// TIA Portal project "XSFW_TIA31001_B0_V15.1" (V15.1)

(* hardware
DEVICE "S7-1200 station_1"  S7-1200 Station
   slot 0: "Rack_0"  S7-1200 Rack  Rack  V1.0
   slot 1: "PLC_Divider"  CPU 1214C DC/DC/DC  6ES7 214-1AG40-0XB0  V4.2
   slot 2: "DI 16/DQ 16x24VDC_1"  6ES7 223-1BL32-0XB0  V2.0
   slot 3: "AI 4x13BIT/AQ 2x14BIT_1"  6ES7 234-4HE32-0XB0  V2.0
   slot 101: "CM 1242-5"  CM 1242-5  6GK7 242-5DX30-0XE0  V1.0
DEVICE "CSM"  SCALANCE X-Station
   slot 0: "Bastidor SCALANCE X"  Rail
   slot 0: "Switch"  6GK7 277-1AA00-0AA0
DEVICE "HMI_1"  KTP700 Basic PN
   slot 0: "HMI_1"  KTP700 Basic PN  6AV2 123-2GB03-0AX0  15.0.0.0
   slot 1: "HMI_RT_1"  KTP700 Basic PN  6AV2 123-2GB03-0AX0  15.0.0.0
   slot 5: "HMI_1.IE_CP_1"  PROFINET Interface  15.0.0.0
      slot 1: "Interfaz PROFINET_1"  PROFINET Interface
         slot 1: "Port_1"  Port
DEVICE "Dispositivo GSD_1"  GSD.Device.PN
   slot 0: "Rack"  Rack  V1.0
   slot 0: "V90-X"  SINAMICS V90 PN V1.0  6SL3 210-5Fxxx-xxFx  V1.00
      slot 0: "SINAMICS V90 PN V1.0"  SINAMICS V90 PN V1.0
      slot 1: "PN-IO"  PN-IO
         slot 1: "Puerto 1"  Port 1
         slot 2: "Puerto 2"  Port 2
      slot 1: "Drive"  Drive
         slot 0: "Punto de acceso a módulo"  Module Access Point
         slot 1: "sin PROFIsafe"  without PROFIsafe
   slot 2: "Telegrama estándar 3, PZD-5/9"  Standard telegram 3, PZD-5/9
DEVICE "Dispositivo GSD_2"  GSD.Device.PN
   slot 0: "Rack"  Rack  V1.0
   slot 0: "V90-Y"  SINAMICS V90 PN V1.0  6SL3 210-5Fxxx-xxFx  V1.00
      slot 0: "SINAMICS V90 PN V1.0"  SINAMICS V90 PN V1.0
      slot 1: "PN-IO"  PN-IO
         slot 1: "Puerto 1"  Port 1
         slot 2: "Puerto 2"  Port 2
      slot 1: "Drive"  Drive
         slot 0: "Punto de acceso a módulo"  Module Access Point
         slot 1: "sin PROFIsafe"  without PROFIsafe
   slot 2: "Telegrama estándar 3, PZD-5/9"  Standard telegram 3, PZD-5/9
*)

// ===== PLC "PLC_Divider"  CPU 1214C DC/DC/DC =====

VAR_GLOBAL   // PLC tag table "Tabla de variables estándar"
   "iCntBot" AT %I0.3 : Bool;
   "iSnsBotBaj" AT %I0.4 : Bool;
   "iSnsBotAlt" AT %I0.5 : Bool;
   "iCH_A" AT %I0.0 : Bool;
   "iCH_B" AT %I0.1 : Bool;
   "iCH_Z" AT %I0.2 : Bool;
   "iSns_Ch1Full" AT %I0.6 : Bool;
   "iSns_Ch2Full" AT %I3.6 : Bool;
   "iSns_Ch3Full" AT %I3.7 : Bool;
   "iSign_HabInv" AT %I3.0 : Bool;
   "iPul_Marcha" AT %I3.1 : Bool;
   "iPul_Parada" AT %I3.2 : Bool;
   "iPul_Rst" AT %I3.3 : Bool;
   "iProt_Abiertas" AT %I3.4 : Bool;
   "iTrip_Inverter" AT %I3.5 : Bool;
   "iRef_Analog" AT %IW54 : Int;
   "qRev_Alarma" AT %Q0.0 : Bool;
   "qSem_Verde" AT %Q0.1 : Bool;
   "qSem_rojo" AT %Q0.2 : Bool;
   "qTest_Marcha" AT %Q0.3 : Bool;
   "qRes_Alarma" AT %Q0.4 : Bool;
   "qRes_Inversor" AT %Q0.5 : Bool;
   "qFwd_Inversor" AT %Q0.6 : Bool;
   "qTrig_2" AT %Q0.7 : Bool;
   "qSign_Marcha" AT %Q1.0 : Bool;
   "qSign_Falla" AT %Q1.1 : Bool;
   "qTrig_1" AT %Q2.0 : Bool;
   "qTrig_22" AT %Q2.1 : Bool;
   "qRef_Analog" AT %IW82 : Int;
   "System_Byte" AT %MB1 : Byte;
   "FirstScan" AT %M1.0 : Bool;
   "DiagStatusUpdate" AT %M1.1 : Bool;
   "AlwaysTRUE" AT %M1.2 : Bool;
   "AlwaysFALSE" AT %M1.3 : Bool;
   "Clock_Byte" AT %MB0 : Byte;
   "Clock_10Hz" AT %M0.0 : Bool;
   "Clock_5Hz" AT %M0.1 : Bool;
   "Clock_2.5Hz" AT %M0.2 : Bool;
   "Clock_2Hz" AT %M0.3 : Bool;
   "Clock_1.25Hz" AT %M0.4 : Bool;
   "Clock_1Hz" AT %M0.5 : Bool;
   "Clock_0.625Hz" AT %M0.6 : Bool;
   "Clock_0.5Hz" AT %M0.7 : Bool;
   "Trip_Inverter" AT %M100.2 : Bool;
   "Marca_Homing" AT %M102.1 : Bool;
   "Eje_X_Drive_IN" AT %I68.0 : "PD_TEL1_IN";
   "Eje_X_Drive_OUT" AT %Q84.0 : "PD_TEL1_OUT";
   "Eje_X_Encoder_IN" AT %I68.0 : "PD_TEL81_IN";
   "Eje_X_Encoder_OUT" AT %Q84.0 : "PD_TEL81_OUT";
   "Eje_Y_Drive_IN" AT %I104.0 : "PD_TEL3_IN";
   "Eje_Y_Drive_OUT" AT %Q74.0 : "PD_TEL3_OUT";
   "Eje_1_Drive_IN" AT %I68.0 : "PD_TEL3_IN";
   "Eje_1_Drive_OUT" AT %Q64.0 : "PD_TEL3_OUT";
   "Tag_1" AT %M102.2 : Bool;
   "MMovX" AT %M850.0 : Bool;
   "Tag_2" AT %M102.3 : Bool;
   "MMovXN" AT %M850.1 : Bool;
   "Tag_3" AT %M102.4 : Bool;
   "MMov2X" AT %M850.2 : Bool;
   "Tag_4" AT %M102.5 : Bool;
   "MMov2XN" AT %M850.3 : Bool;
   "Tag_5" AT %M102.6 : Bool;
   "MMovY" AT %M850.4 : Bool;
   "MMovYN" AT %M850.5 : Bool;
   "Tag_6" AT %M102.7 : Bool;
   "Eje_Y_Drive_IN(1)" AT %I86.0 : "PD_TEL3_IN";
   "Tag_7" AT %M110.0 : Bool;
   "Tag_8" AT %M110.1 : Bool;
   "Tag_9" AT %M110.2 : Bool;
   "Tag_10" AT %M110.3 : Bool;
   "Tag_11" AT %M110.4 : Bool;
   "Tag_12" AT %M110.5 : Bool;
   "Tag_13" AT %M800.1 : Bool;
   "Tag_14" AT %M103.0 : Bool;
   "Tag_15" AT %M103.1 : Bool;
   "Tag_16" AT %M1000.0 : Bool;
   "iHsc_Z" AT %ID1000 : DInt;
   "Hsc_Za" AT %MD20 : DInt;
   "iPulsos0.1Seg" AT %MD24 : DInt;
   "Contando" AT %M150.0 : Bool;
   "Fin_Cuenta" AT %M150.1 : Bool;
   "Halt_Motor" AT %M150.2 : Bool;
   "Band_E24" AT %M150.3 : Bool;
   "Tag_17" AT %M800.0 : Bool;
   "Band_E22" AT %M150.4 : Bool;
   "Band_E23" AT %M150.5 : Bool;
   "Tag_18" AT %MD22 : DInt;
   "Hsc_Zb" AT %MD28 : DInt;
   "Hsc_sub" AT %MD32 : DInt;
   "Hsc_sub1" AT %MD36 : DInt;
   "Error_Velocidad" AT %M150.6 : Bool;
   "Enc_hab" AT %E104.0 : Bool;
   "Enc_stop" AT %I104.1 : Bool;
   "Tag_19" AT %IW104 : Word;
   "Tag_20" AT %IW106 : Word;
   "Tag_21" AT %IW108 : Word;
   "Tag_22" AT %IW110 : Word;
   "Tag_23" AT %QW104 : Word;
   "Tag_24" AT %QW106 : Word;
   "Tag_25" AT %QW108 : Word;
   "Tag_26" AT %QW110 : Word;
END_VAR

VAR_GLOBAL   // PLC tag table "Alarmas"
   "Alarmas_1" AT %MW100 : Word;
   "ProteccionAbierta" AT %M100.0 : Bool;   // Señal I3.4 en 1
   "BotellaCaida" AT %M100.1 : Bool;
END_VAR

VAR_GLOBAL   // PLC tag table "Inicializaciòn"
   "Marcas para la inicializaciòn" AT %MW102 : Word;
   "Start" AT %M102.0 : Bool;
END_VAR

DATA_BLOCK "01_LINEA_Entradas-DB"   // DB1
{ S7_Optimized_Access := 'TRUE' }
VERSION : 0.1
   VAR
      Contador : Bool;   // Pulsador de marcha
      Sensor_Bajo : Bool;   // Pulsador de parada
      Sensor_Alto : Bool;   // Pulsador de marcha columna 4
      CH_A : Bool;   // Pulsador de parada de emergancia columna 4
      CH_B : Bool;   // Pulsador de marcha columna 6
      CH_Z : Bool;   // Pulsador de parada de emergancia columna 6
      Canal1_Full : Bool;   // Pulsador de marcha columna 9
      Canal2_Full : Bool;   // Pulsador de parada de emergancia columna 9
      Canal3_Full : Bool;   // Pulsador de marcha columna 11
      Hab_Inverter : Bool;   // Pulsador de parada de emergancia columna 11
      Marcha : Bool;   // Pulsador de marcha columna 12
      Parada : Bool;   // Pulsador de parada de emergancia columna 12
      Reset : Bool;   // Pulsador de parada de emergancia del tablero general
      Protecciones_Abiertas : Bool;   // Pulsador de parada de emergencia del tablero de la fosa
      Trip_Inverter : Bool;   // Señal de falla del variador
      Enc_andando : Bool;
      Enc_parada : Bool;
   END_VAR
BEGIN
END_DATA_BLOCK

DATA_BLOCK "02_LINEA_Salidas-DB"   // DB2
{ S7_Optimized_Access := 'TRUE' }
VERSION : 0.1
   VAR
      Alarma_Sonora : Bool;   // Marcha para el variador
      Semaforo_Verde : Bool;   // Sentido adelante variador
      Semaforo_Rojo : Bool;   // Sentido atras variador
      Testigo_Marcha : Bool;   // Indicador sonoro
      Reset_Alarma : Bool;   // Indicador de linea en marcha
      Reset_Inverter : Bool;   // Indicador de linea parada
      Avance_Inverter : Bool;   // Buzzer de la baliza del tablero principal
      Trigger_2 : Bool;   // Lampara verde de la baliza del tablero principal
      EnMarcha : Bool;   // Lampara roja de la baliza del tablero principal
      EnFalla : Bool;   // Lampara amarilla de la baliza del tablero principal
      Trigger_11 : Bool;
      Trigger_22 : Bool;
      Ref_20mA : Int;
   END_VAR
BEGIN
END_DATA_BLOCK

DATA_BLOCK "MotorInverter"   // DB5
{ S7_Optimized_Access := 'TRUE' }
VERSION : 0.1
// stored: InstanceOfName Motor Simple
"Motor Simple"
BEGIN
END_DATA_BLOCK

DATA_BLOCK "FB_INC_GENERAL_DB"   // DB7
{ S7_Optimized_Access := 'FALSE' }
VERSION : 0.1
// stored: InstanceOfName FB_INC_GENERAL
"FB_INC_GENERAL"
BEGIN
END_DATA_BLOCK

DATA_BLOCK "Cuentas_Matematicas1_DB"   // DB15
{ S7_Optimized_Access := 'TRUE' }
VERSION : 0.1
   VAR
      MovXNeg : Real := 0.0;
      Mov2X : Real := 0.0;
      Mov2XNeg : Real := 0.0;
      MovYNeg : Real := 0.0;
   END_VAR
BEGIN
END_DATA_BLOCK

DATA_BLOCK "FB_GENERAL_DB"   // DB17
{ S7_Optimized_Access := 'FALSE' }
VERSION : 0.1
// stored: InstanceOfName FB_GENERAL
"FB_GENERAL"
BEGIN
END_DATA_BLOCK

DATA_BLOCK "Cuentas_Matematicas1_DB_1"   // DB20
{ S7_Optimized_Access := 'TRUE' }
VERSION : 0.1
// stored: InstanceOfName Cuentas_Matematicas1
"Cuentas_Matematicas1"
BEGIN
END_DATA_BLOCK

DATA_BLOCK "DB_Encajonadora"   // DB28
{ S7_Optimized_Access := 'TRUE' }
VERSION : 0.1
   VAR
      Word1 : Word;   // bit 0 y 1 para guardar estado de encajonadora
      Word2 : Word;
      Word3 : Word;
      Word4 : Word;
      Word5 : Word;
      Word6 : Word;
      Word7 : Word;
      Word8 : Word;
   END_VAR
BEGIN
END_DATA_BLOCK

DATA_BLOCK "DB_GENERAL"   // DB100
{ S7_Optimized_Access := 'FALSE' }
VERSION : 0.1
// stored: InstanceOfName FB_GENERAL
"FB_GENERAL"
BEGIN
END_DATA_BLOCK

// folder: COMANDOS

DATA_BLOCK "DB_SUB_0_COM_GENERAL"   // DB600
{ S7_Optimized_Access := 'FALSE' }
VERSION : 0.1
   VAR
      ManipEsperaCarro : Bool;
      RecepCarroConfir : Bool;
      SalidaEsperaCarro1 : Bool;
      SalidaEsperaCarro2 : Bool;
      TengoCarroEnPortacarro : Bool;
      ReconocimientoAlarmas : Bool;
   END_VAR
BEGIN
END_DATA_BLOCK

// folder: INCIDENTES

DATA_BLOCK "DB_INC_GENERAL"   // DB500
{ S7_Optimized_Access := 'FALSE' }
VERSION : 0.1
// stored: InstanceOfName FB_INC_GENERAL
"FB_INC_GENERAL"
BEGIN
END_DATA_BLOCK

// folder: PUESTA EN MARCHA

DATA_BLOCK "DB_PUESTA_MARCHA"   // DB10
{ S7_Optimized_Access := 'TRUE' }
VERSION : 0.1
   VAR RETAIN
      MovYmm : Real := 30.0;
      MovXmm : Real := 30.0;
   END_VAR
   VAR
      TChFull : Time := T#1S;
   END_VAR
BEGIN
END_DATA_BLOCK

// folder: System blocks/Program resources

DATA_BLOCK "IEC_Counter_0_DB"   // DB6
{ S7_Optimized_Access := 'TRUE' }
AUTHOR : Simatic
FAMILY : IEC
NAME : CNTR
VERSION : 1.0
// stored: InstanceOfName IEC_COUNTER
"IEC_COUNTER"
BEGIN
END_DATA_BLOCK

DATA_BLOCK "IEC_Counter_1_DB"   // DB8
{ S7_Optimized_Access := 'TRUE' }
AUTHOR : Simatic
FAMILY : IEC
NAME : CNTR
VERSION : 1.0
// stored: InstanceOfName IEC_COUNTER
"IEC_COUNTER"
BEGIN
END_DATA_BLOCK

DATA_BLOCK "IEC_Counter_2_DB"   // DB9
{ S7_Optimized_Access := 'TRUE' }
AUTHOR : Simatic
FAMILY : IEC
NAME : CNTR
VERSION : 1.0
// stored: InstanceOfName IEC_COUNTER
"IEC_COUNTER"
BEGIN
END_DATA_BLOCK

DATA_BLOCK "IEC_Timer_ChFull"   // DB11
{ S7_Optimized_Access := 'TRUE' }
AUTHOR : Simatic
FAMILY : IEC
NAME : IEC_TMR
VERSION : 1.0
// stored: InstanceOfName IEC_TIMER
"IEC_TIMER"
BEGIN
END_DATA_BLOCK

DATA_BLOCK "IEC_Timer_0_DB_1"   // DB30
{ S7_Optimized_Access := 'TRUE' }
AUTHOR : Simatic
FAMILY : IEC
NAME : IEC_TMR
VERSION : 1.0
// stored: InstanceOfName IEC_TIMER
"IEC_TIMER"
BEGIN
END_DATA_BLOCK

DATA_BLOCK "IEC_Timer_0_DB_2"   // DB31
{ S7_Optimized_Access := 'TRUE' }
AUTHOR : Simatic
FAMILY : IEC
NAME : IEC_TMR
VERSION : 1.0
// stored: InstanceOfName IEC_TIMER
"IEC_TIMER"
BEGIN
END_DATA_BLOCK

DATA_BLOCK "IEC_Timer_0_DB_3"   // DB32
{ S7_Optimized_Access := 'TRUE' }
AUTHOR : Simatic
FAMILY : IEC
NAME : IEC_TMR
VERSION : 1.0
// stored: InstanceOfName IEC_TIMER
"IEC_TIMER"
BEGIN
END_DATA_BLOCK

DATA_BLOCK "IEC_Timer_0_DB_4"   // DB33
{ S7_Optimized_Access := 'TRUE' }
AUTHOR : Simatic
FAMILY : IEC
NAME : IEC_TMR
VERSION : 1.0
// stored: InstanceOfName IEC_TIMER
"IEC_TIMER"
BEGIN
END_DATA_BLOCK

DATA_BLOCK "IEC_Timer_0_DB_5"   // DB34
{ S7_Optimized_Access := 'TRUE' }
AUTHOR : Simatic
FAMILY : IEC
NAME : IEC_TMR
VERSION : 1.0
// stored: InstanceOfName IEC_TIMER
"IEC_TIMER"
BEGIN
END_DATA_BLOCK

// folder: VISUALIZACION

DATA_BLOCK "DB_VIS_GENERAL"   // DB800
{ S7_Optimized_Access := 'FALSE' }
VERSION : 0.1
   VAR
      CantBot : Int;
      AlarmaProtecciòn : Bool;
      AlarmaBotellaCaida : Bool;
      MC_Pwr_EnX : Bool;
      MC_Pwrt_EnY : Bool;
      MC_Res_ExX : Bool;
      MC_Res_ExY : Bool;
      MC_JogFwd_X : Bool;
      MC_JogFwd_Y : Bool;
      MC_JogBwd_X : Bool;
      MC_JogBwd_Y : Bool;
      HomingOk : Bool;
      Reset : Bool;
      Start : Bool;
   END_VAR
BEGIN
END_DATA_BLOCK

// folder: (top level)

DATA_BLOCK "Eje_Y"   // DB4, Motion_DB
{ S7_Optimized_Access := 'TRUE' }
AUTHOR : SIMATIC
FAMILY : BasicMC
NAME : TO_PosAx
VERSION : 6.0
// stored: InstanceOfName TO_PositioningAxis
"TO_PositioningAxis"
BEGIN
   // Axis.Encoder.TelegramAddressOutCU = %Q74.0
   // Axis.Encoder.TelegramAddressInCU = %I86.0
   // Axis.Encoder.DoNameCU = V90-Y.Drive_Encóder1
   // Axis.Drive.TelegramAddressOutCU = %Q74.0
   // Axis.Drive.TelegramAddressInCU = %I86.0
   // Axis.Drive.TelegramType = 2
   // Axis.Drive.DoNameCU = V90-Y.Drive
   // Axis.LengthUnitNormalized.Time = 1
   // Axis.LengthUnitNormalized.Distance = -2
   // Axis.Encoder.SelectedHscIndexCU = -1
   // Axis.Encoder.DbTypeCU = Classic
   // Axis.Drive.DbTypeCU = Classic
END_DATA_BLOCK

DATA_BLOCK "Eje_X"   // DB12, Motion_DB
{ S7_Optimized_Access := 'TRUE' }
AUTHOR : SIMATIC
FAMILY : BasicMC
NAME : TO_PosAx
VERSION : 6.0
// stored: InstanceOfName TO_PositioningAxis
"TO_PositioningAxis"
BEGIN
   // Axis.Encoder.TelegramAddressOutCU = %Q64.0
   // Axis.Encoder.TelegramAddressInCU = %I68.0
   // Axis.Encoder.DoNameCU = V90-X.Drive_Encóder1
   // Axis.Drive.TelegramAddressOutCU = %Q64.0
   // Axis.Drive.TelegramAddressInCU = %I68.0
   // Axis.Drive.TelegramType = 2
   // Axis.Drive.DoNameCU = V90-X.Drive
   // Axis.LengthUnitNormalized.Distance = 1013
   // Axis.Encoder.SelectedHscIndexCU = -1
   // Axis.Encoder.DbTypeCU = Classic
   // Axis.Drive.DbTypeCU = Classic
END_DATA_BLOCK

FUNCTION_BLOCK "Cuentas_Matematicas1"   // FB1, LAD
TITLE = ---------------------------Calculo de distancias----------------------------------------
{ S7_Optimized_Access := 'TRUE' }
VERSION : 0.1
BEGIN

REGION Network 1: Movimiento negativo en X
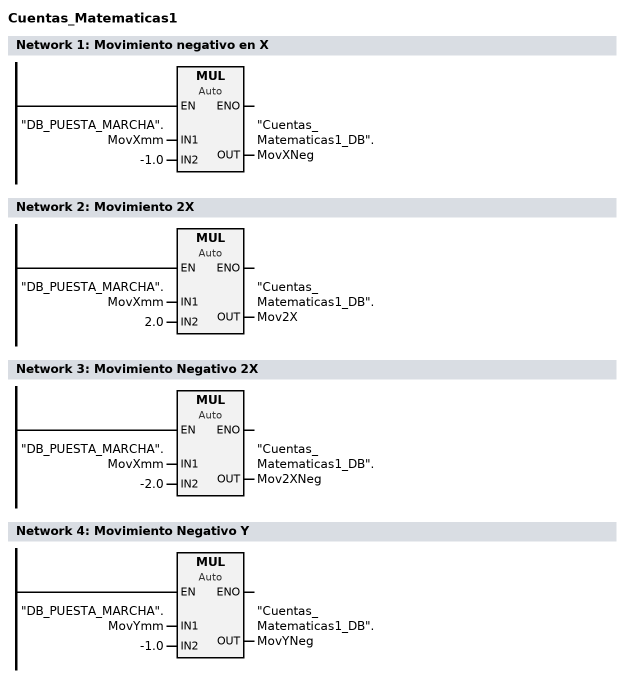
   RUNG wire#powerrail
      Mul(in1 := "DB_PUESTA_MARCHA".MovXmm, in2 := -1.0, out => "Cuentas_Matematicas1_DB".MovXNeg)
   END_RUNG
   // the same network as SCL:
   "Cuentas_Matematicas1_DB".MovXNeg := "DB_PUESTA_MARCHA".MovXmm * (-1.0);
END_REGION

REGION Network 2: Movimiento 2X
   RUNG wire#powerrail
      Mul(in1 := "DB_PUESTA_MARCHA".MovXmm, in2 := 2.0, out => "Cuentas_Matematicas1_DB".Mov2X)
   END_RUNG
   // the same network as SCL:
   "Cuentas_Matematicas1_DB".Mov2X := "DB_PUESTA_MARCHA".MovXmm * 2.0;
END_REGION

REGION Network 3: Movimiento Negativo 2X
   RUNG wire#powerrail
      Mul(in1 := "DB_PUESTA_MARCHA".MovXmm, in2 := -2.0, out => "Cuentas_Matematicas1_DB".Mov2XNeg)
   END_RUNG
   // the same network as SCL:
   "Cuentas_Matematicas1_DB".Mov2XNeg := "DB_PUESTA_MARCHA".MovXmm * (-2.0);
END_REGION

REGION Network 4: Movimiento Negativo Y
   RUNG wire#powerrail
      Mul(in1 := "DB_PUESTA_MARCHA".MovYmm, in2 := -1.0, out => "Cuentas_Matematicas1_DB".MovYNeg)
   END_RUNG
   // the same network as SCL:
   "Cuentas_Matematicas1_DB".MovYNeg := "DB_PUESTA_MARCHA".MovYmm * (-1.0);
END_REGION
END_FUNCTION_BLOCK

FUNCTION_BLOCK "FB_GENERAL"   // FB100, LAD
{ S7_Optimized_Access := 'FALSE' }
VERSION : 0.1
   VAR_OUTPUT
      DoneX : Bool;
      DoneXN : Bool;
      DoneY : Bool;
      DoneYN : Bool;
      Done2X : Bool;
      Done2XN : Bool;
   END_VAR
   VAR
      Estados : Array[0..32] of Bool;
      Concatenadoras : Array[0..32] of Bool;
      Prioritarias : Array[0..32] of Bool;
      Error_Concatenadoras : Bool;
      Error_Prioritarias : Bool;
      Cuenta_1 : Bool;
      Cuenta_2 : Bool;
      Cuenta_3 : Bool;
      "Cont_Botellas/2" : Int;
   END_VAR
BEGIN

REGION Network 1: Inicializaciòn
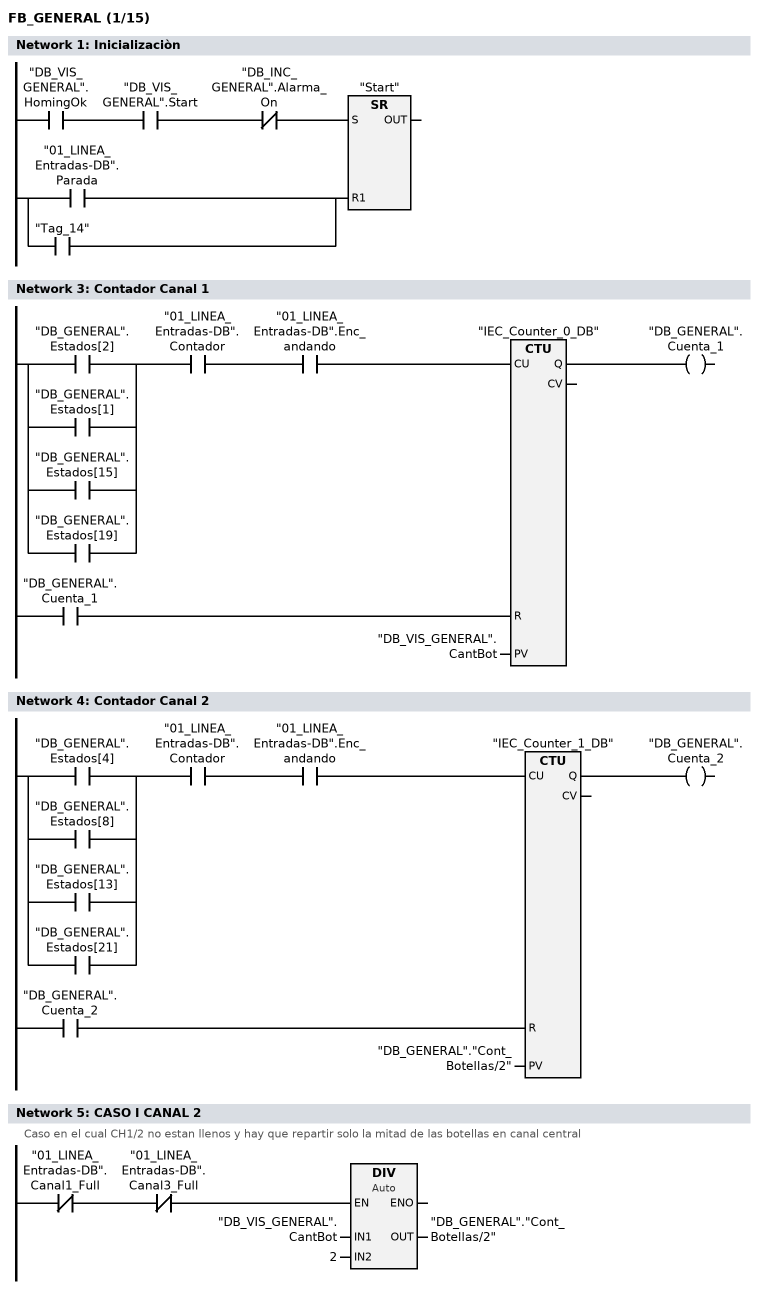
   RUNG wire#powerrail
      Contact( "DB_VIS_GENERAL".HomingOk )
      Contact( "DB_VIS_GENERAL".Start )
      I_Contact( "DB_INC_GENERAL".Alarma_On )
      S_SR(operand := "Start", r1 := wire#w1)
   END_RUNG
   RUNG wire#powerrail
      Contact( "01_LINEA_Entradas-DB".Parada )
   END_RUNG wire#w1
   RUNG wire#powerrail
      Contact( "Tag_14" )
   END_RUNG wire#w1
   // the same network as SCL:
   IF "DB_VIS_GENERAL".HomingOk AND "DB_VIS_GENERAL".Start AND NOT "DB_INC_GENERAL".Alarma_On THEN
       "Start" := TRUE;   // SR flip-flop
   END_IF;
   IF "01_LINEA_Entradas-DB".Parada OR "Tag_14" THEN "Start" := FALSE; END_IF;
END_REGION

REGION Network 2: -----------------OTROS---------------
END_REGION

REGION Network 3: Contador Canal 1
   "IEC_Counter_0_DB".CTU(CU := ("DB_GENERAL".Estados[2] OR "DB_GENERAL".Estados[1] OR "DB_GENERAL".Estados[15] OR "DB_GENERAL".Estados[19]) AND "01_LINEA_Entradas-DB".Contador AND "01_LINEA_Entradas-DB".Enc_andando,
                          R := "DB_GENERAL".Cuenta_1,
                          PV := "DB_VIS_GENERAL".CantBot);
   "DB_GENERAL".Cuenta_1 := "IEC_Counter_0_DB".Q;
END_REGION

REGION Network 4: Contador Canal 2
   "IEC_Counter_1_DB".CTU(CU := ("DB_GENERAL".Estados[4] OR "DB_GENERAL".Estados[8] OR "DB_GENERAL".Estados[13] OR "DB_GENERAL".Estados[21]) AND "01_LINEA_Entradas-DB".Contador AND "01_LINEA_Entradas-DB".Enc_andando,
                          R := "DB_GENERAL".Cuenta_2,
                          PV := "DB_GENERAL"."Cont_Botellas/2");
   "DB_GENERAL".Cuenta_2 := "IEC_Counter_1_DB".Q;
END_REGION

REGION Network 5: CASO I CANAL 2
   // Caso en el cual CH1/2 no estan llenos y hay que repartir solo la mitad de las botellas en canal central
   RUNG wire#powerrail
      I_Contact( "01_LINEA_Entradas-DB".Canal1_Full )
      I_Contact( "01_LINEA_Entradas-DB".Canal3_Full )
      Div(in1 := "DB_VIS_GENERAL".CantBot, in2 := 2, out => "DB_GENERAL"."Cont_Botellas/2")
   END_RUNG
   // the same network as SCL:
   IF NOT "01_LINEA_Entradas-DB".Canal1_Full AND NOT "01_LINEA_Entradas-DB".Canal3_Full THEN
       "DB_GENERAL"."Cont_Botellas/2" := "DB_VIS_GENERAL".CantBot / 2;
   END_IF;
END_REGION

REGION Network 6: CASO II CANAL 2
   // Caso en el cual CH1/2 estan llenos y hay que repartir la misma cantidad de botellas en el carril central.
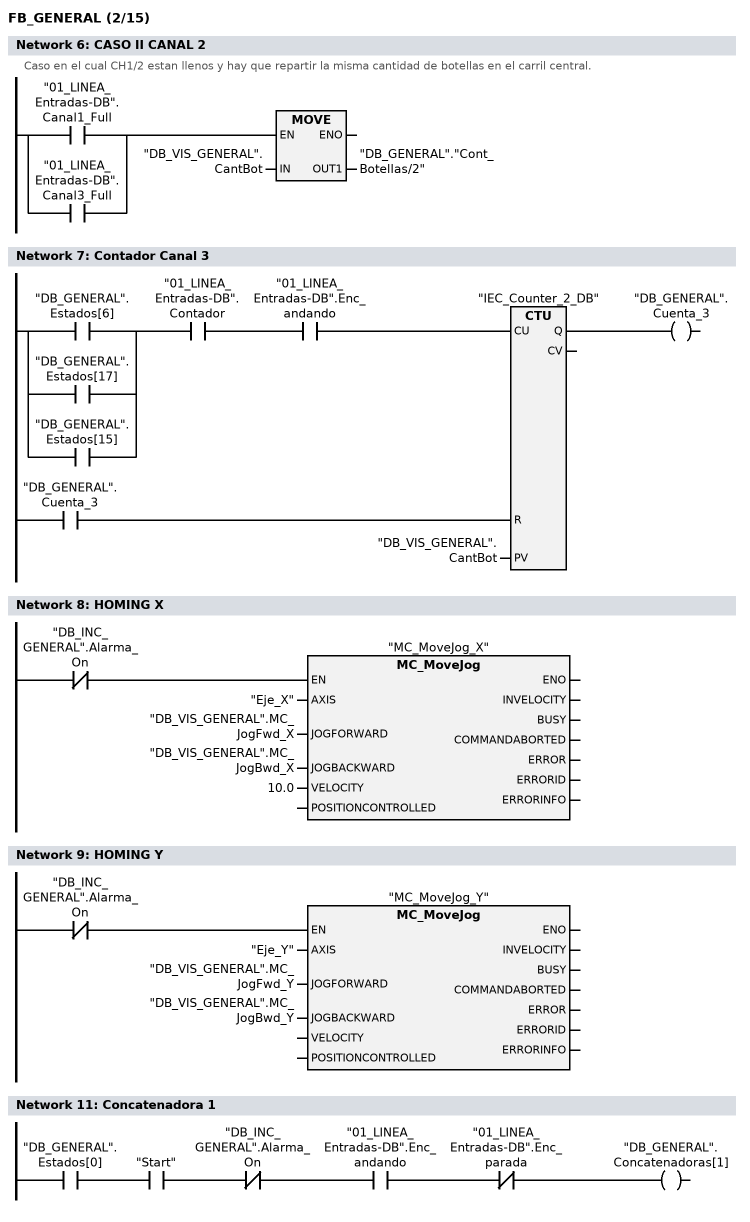
   RUNG wire#powerrail
      Contact( "01_LINEA_Entradas-DB".Canal1_Full )
      wire#w1
      Move(in := "DB_VIS_GENERAL".CantBot, out1 => "DB_GENERAL"."Cont_Botellas/2")
   END_RUNG
   RUNG wire#powerrail
      Contact( "01_LINEA_Entradas-DB".Canal3_Full )
   END_RUNG wire#w1
   // the same network as SCL:
   IF "01_LINEA_Entradas-DB".Canal1_Full OR "01_LINEA_Entradas-DB".Canal3_Full THEN
       "DB_GENERAL"."Cont_Botellas/2" := "DB_VIS_GENERAL".CantBot;
   END_IF;
END_REGION

REGION Network 7: Contador Canal 3
   "IEC_Counter_2_DB".CTU(CU := ("DB_GENERAL".Estados[6] OR "DB_GENERAL".Estados[17] OR "DB_GENERAL".Estados[15]) AND "01_LINEA_Entradas-DB".Contador AND "01_LINEA_Entradas-DB".Enc_andando,
                          R := "DB_GENERAL".Cuenta_3,
                          PV := "DB_VIS_GENERAL".CantBot);
   "DB_GENERAL".Cuenta_3 := "IEC_Counter_2_DB".Q;
END_REGION

REGION Network 8: HOMING X
   IF NOT "DB_INC_GENERAL".Alarma_On THEN
       "MC_MoveJog_X"(Axis := "Eje_X",   // MC_MoveJog
                      JogForward := "DB_VIS_GENERAL".MC_JogFwd_X,
                      JogBackward := "DB_VIS_GENERAL".MC_JogBwd_X,
                      Velocity := 10.0);
   END_IF;
END_REGION

REGION Network 9: HOMING Y
   IF NOT "DB_INC_GENERAL".Alarma_On THEN
       "MC_MoveJog_Y"(Axis := "Eje_Y",   // MC_MoveJog
                      JogForward := "DB_VIS_GENERAL".MC_JogFwd_Y,
                      JogBackward := "DB_VIS_GENERAL".MC_JogBwd_Y);
   END_IF;
END_REGION

REGION Network 10: --------------------Maquina de estados - 3 carriles-----------------
END_REGION

REGION Network 11: Concatenadora 1
   RUNG wire#powerrail
      Contact( "DB_GENERAL".Estados[0] )
      Contact( "Start" )
      I_Contact( "DB_INC_GENERAL".Alarma_On )
      Contact( "01_LINEA_Entradas-DB".Enc_andando )
      I_Contact( "01_LINEA_Entradas-DB".Enc_parada )
      Coil( "DB_GENERAL".Concatenadoras[1] )
   END_RUNG
   // the same network as SCL:
   "DB_GENERAL".Concatenadoras[1] := "DB_GENERAL".Estados[0] AND "Start" AND NOT "DB_INC_GENERAL".Alarma_On AND "01_LINEA_Entradas-DB".Enc_andando AND NOT "01_LINEA_Entradas-DB".Enc_parada;
END_REGION

REGION Network 12: Concatenadora 2 (3)
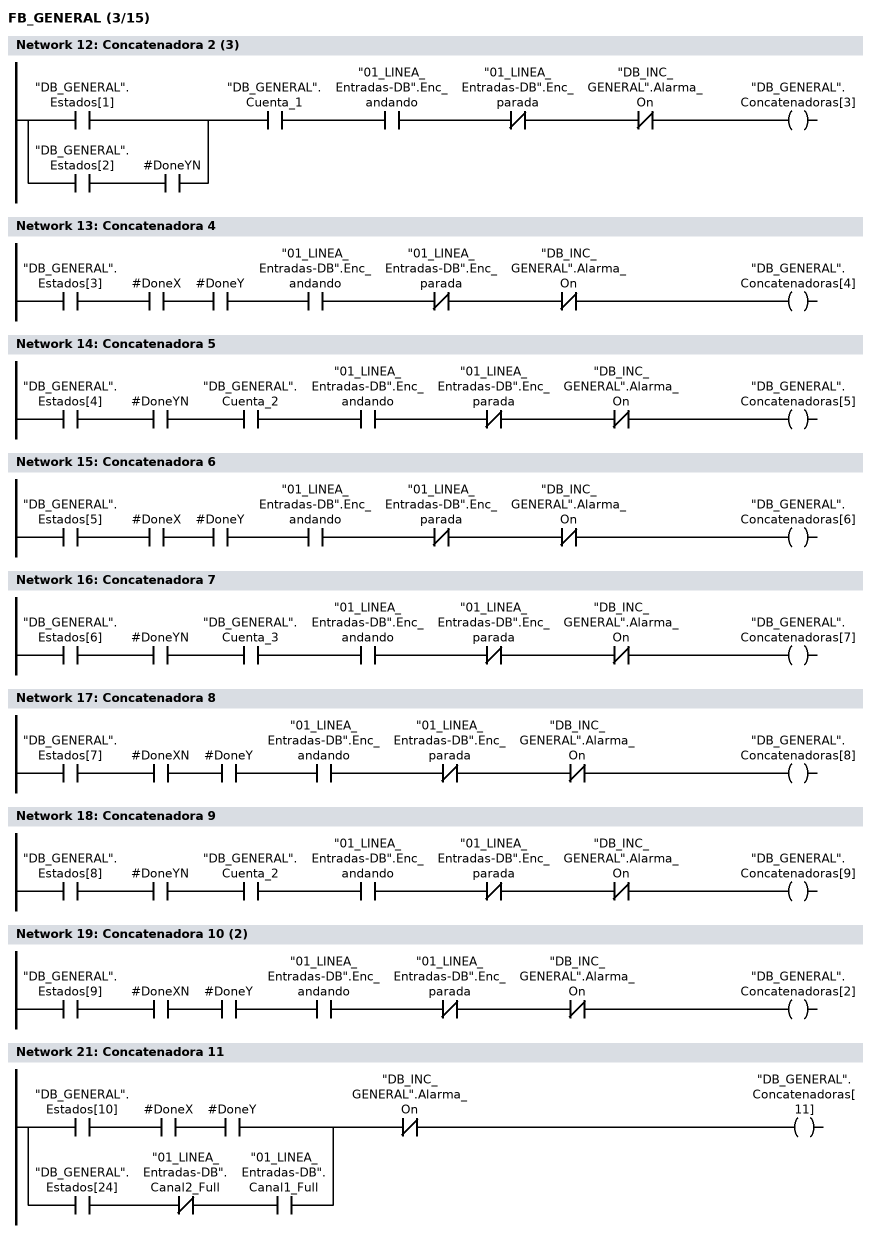
   RUNG wire#powerrail
      Contact( "DB_GENERAL".Estados[1] )
      wire#w1
      Contact( "DB_GENERAL".Cuenta_1 )
      Contact( "01_LINEA_Entradas-DB".Enc_andando )
      I_Contact( "01_LINEA_Entradas-DB".Enc_parada )
      I_Contact( "DB_INC_GENERAL".Alarma_On )
      Coil( "DB_GENERAL".Concatenadoras[3] )
   END_RUNG
   RUNG wire#powerrail
      Contact( "DB_GENERAL".Estados[2] )
      Contact( #DoneYN )
   END_RUNG wire#w1
   // the same network as SCL:
   "DB_GENERAL".Concatenadoras[3] := ("DB_GENERAL".Estados[1] OR ("DB_GENERAL".Estados[2] AND #DoneYN)) AND "DB_GENERAL".Cuenta_1 AND "01_LINEA_Entradas-DB".Enc_andando AND NOT "01_LINEA_Entradas-DB".Enc_parada AND NOT "DB_INC_GENERAL".Alarma_On;
END_REGION

REGION Network 13: Concatenadora 4
   RUNG wire#powerrail
      Contact( "DB_GENERAL".Estados[3] )
      Contact( #DoneX )
      Contact( #DoneY )
      Contact( "01_LINEA_Entradas-DB".Enc_andando )
      I_Contact( "01_LINEA_Entradas-DB".Enc_parada )
      I_Contact( "DB_INC_GENERAL".Alarma_On )
      Coil( "DB_GENERAL".Concatenadoras[4] )
   END_RUNG
   // the same network as SCL:
   "DB_GENERAL".Concatenadoras[4] := "DB_GENERAL".Estados[3] AND #DoneX AND #DoneY AND "01_LINEA_Entradas-DB".Enc_andando AND NOT "01_LINEA_Entradas-DB".Enc_parada AND NOT "DB_INC_GENERAL".Alarma_On;
END_REGION

REGION Network 14: Concatenadora 5
   RUNG wire#powerrail
      Contact( "DB_GENERAL".Estados[4] )
      Contact( #DoneYN )
      Contact( "DB_GENERAL".Cuenta_2 )
      Contact( "01_LINEA_Entradas-DB".Enc_andando )
      I_Contact( "01_LINEA_Entradas-DB".Enc_parada )
      I_Contact( "DB_INC_GENERAL".Alarma_On )
      Coil( "DB_GENERAL".Concatenadoras[5] )
   END_RUNG
   // the same network as SCL:
   "DB_GENERAL".Concatenadoras[5] := "DB_GENERAL".Estados[4] AND #DoneYN AND "DB_GENERAL".Cuenta_2 AND "01_LINEA_Entradas-DB".Enc_andando AND NOT "01_LINEA_Entradas-DB".Enc_parada AND NOT "DB_INC_GENERAL".Alarma_On;
END_REGION

REGION Network 15: Concatenadora 6
   RUNG wire#powerrail
      Contact( "DB_GENERAL".Estados[5] )
      Contact( #DoneX )
      Contact( #DoneY )
      Contact( "01_LINEA_Entradas-DB".Enc_andando )
      I_Contact( "01_LINEA_Entradas-DB".Enc_parada )
      I_Contact( "DB_INC_GENERAL".Alarma_On )
      Coil( "DB_GENERAL".Concatenadoras[6] )
   END_RUNG
   // the same network as SCL:
   "DB_GENERAL".Concatenadoras[6] := "DB_GENERAL".Estados[5] AND #DoneX AND #DoneY AND "01_LINEA_Entradas-DB".Enc_andando AND NOT "01_LINEA_Entradas-DB".Enc_parada AND NOT "DB_INC_GENERAL".Alarma_On;
END_REGION

REGION Network 16: Concatenadora 7
   RUNG wire#powerrail
      Contact( "DB_GENERAL".Estados[6] )
      Contact( #DoneYN )
      Contact( "DB_GENERAL".Cuenta_3 )
      Contact( "01_LINEA_Entradas-DB".Enc_andando )
      I_Contact( "01_LINEA_Entradas-DB".Enc_parada )
      I_Contact( "DB_INC_GENERAL".Alarma_On )
      Coil( "DB_GENERAL".Concatenadoras[7] )
   END_RUNG
   // the same network as SCL:
   "DB_GENERAL".Concatenadoras[7] := "DB_GENERAL".Estados[6] AND #DoneYN AND "DB_GENERAL".Cuenta_3 AND "01_LINEA_Entradas-DB".Enc_andando AND NOT "01_LINEA_Entradas-DB".Enc_parada AND NOT "DB_INC_GENERAL".Alarma_On;
END_REGION

REGION Network 17: Concatenadora 8
   RUNG wire#powerrail
      Contact( "DB_GENERAL".Estados[7] )
      Contact( #DoneXN )
      Contact( #DoneY )
      Contact( "01_LINEA_Entradas-DB".Enc_andando )
      I_Contact( "01_LINEA_Entradas-DB".Enc_parada )
      I_Contact( "DB_INC_GENERAL".Alarma_On )
      Coil( "DB_GENERAL".Concatenadoras[8] )
   END_RUNG
   // the same network as SCL:
   "DB_GENERAL".Concatenadoras[8] := "DB_GENERAL".Estados[7] AND #DoneXN AND #DoneY AND "01_LINEA_Entradas-DB".Enc_andando AND NOT "01_LINEA_Entradas-DB".Enc_parada AND NOT "DB_INC_GENERAL".Alarma_On;
END_REGION

REGION Network 18: Concatenadora 9
   RUNG wire#powerrail
      Contact( "DB_GENERAL".Estados[8] )
      Contact( #DoneYN )
      Contact( "DB_GENERAL".Cuenta_2 )
      Contact( "01_LINEA_Entradas-DB".Enc_andando )
      I_Contact( "01_LINEA_Entradas-DB".Enc_parada )
      I_Contact( "DB_INC_GENERAL".Alarma_On )
      Coil( "DB_GENERAL".Concatenadoras[9] )
   END_RUNG
   // the same network as SCL:
   "DB_GENERAL".Concatenadoras[9] := "DB_GENERAL".Estados[8] AND #DoneYN AND "DB_GENERAL".Cuenta_2 AND "01_LINEA_Entradas-DB".Enc_andando AND NOT "01_LINEA_Entradas-DB".Enc_parada AND NOT "DB_INC_GENERAL".Alarma_On;
END_REGION

REGION Network 19: Concatenadora 10 (2)
   RUNG wire#powerrail
      Contact( "DB_GENERAL".Estados[9] )
      Contact( #DoneXN )
      Contact( #DoneY )
      Contact( "01_LINEA_Entradas-DB".Enc_andando )
      I_Contact( "01_LINEA_Entradas-DB".Enc_parada )
      I_Contact( "DB_INC_GENERAL".Alarma_On )
      Coil( "DB_GENERAL".Concatenadoras[2] )
   END_RUNG
   // the same network as SCL:
   "DB_GENERAL".Concatenadoras[2] := "DB_GENERAL".Estados[9] AND #DoneXN AND #DoneY AND "01_LINEA_Entradas-DB".Enc_andando AND NOT "01_LINEA_Entradas-DB".Enc_parada AND NOT "DB_INC_GENERAL".Alarma_On;
END_REGION

REGION Network 20: ---------------Maquina de estado - 2 carriles -------------
END_REGION

REGION Network 21: Concatenadora 11
   RUNG wire#powerrail
      Contact( "DB_GENERAL".Estados[10] )
      Contact( #DoneX )
      Contact( #DoneY )
      wire#w1
      I_Contact( "DB_INC_GENERAL".Alarma_On )
      Coil( "DB_GENERAL".Concatenadoras[11] )
   END_RUNG
   RUNG wire#powerrail
      Contact( "DB_GENERAL".Estados[24] )
      I_Contact( "01_LINEA_Entradas-DB".Canal2_Full )
      Contact( "01_LINEA_Entradas-DB".Canal1_Full )
   END_RUNG wire#w1
   // the same network as SCL:
   "DB_GENERAL".Concatenadoras[11] := (("DB_GENERAL".Estados[10] AND #DoneX AND #DoneY) OR ("DB_GENERAL".Estados[24] AND NOT "01_LINEA_Entradas-DB".Canal2_Full AND "01_LINEA_Entradas-DB".Canal1_Full)) AND NOT "DB_INC_GENERAL".Alarma_On;
END_REGION

REGION Network 22: Concatenadora 12
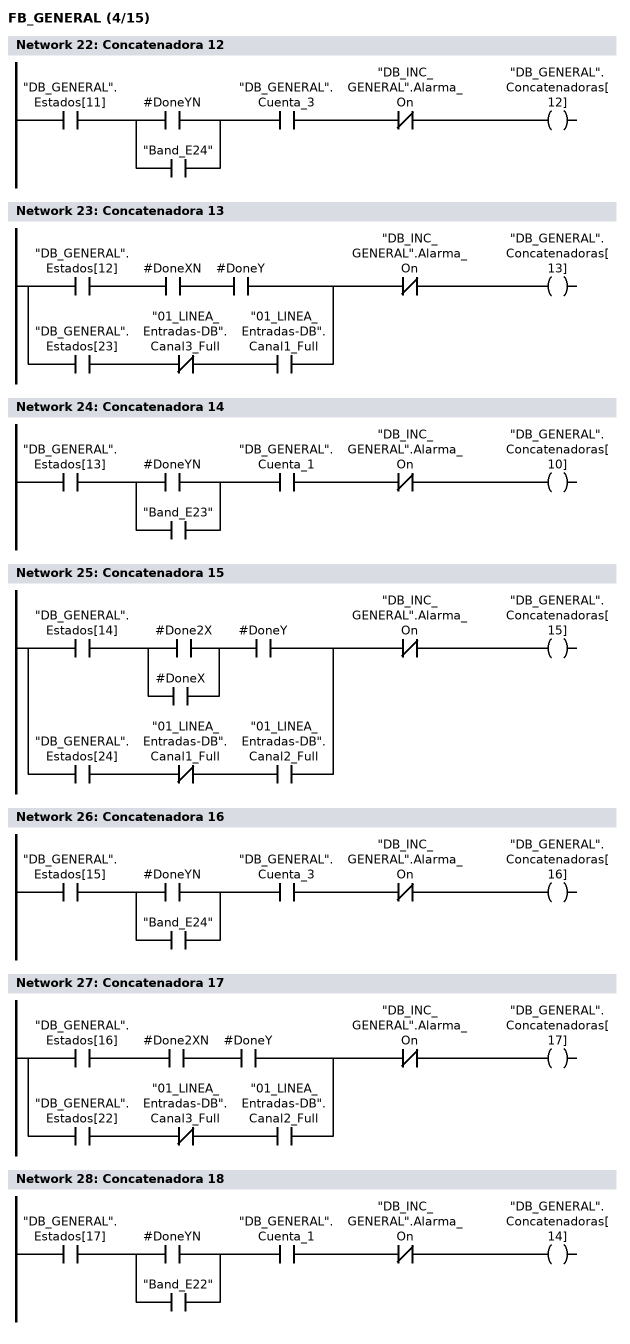
   RUNG wire#powerrail
      Contact( "DB_GENERAL".Estados[11] )
      wire#w1
      Contact( #DoneYN )
      wire#w2
      Contact( "DB_GENERAL".Cuenta_3 )
      I_Contact( "DB_INC_GENERAL".Alarma_On )
      Coil( "DB_GENERAL".Concatenadoras[12] )
   END_RUNG
   RUNG wire#w1
      Contact( "Band_E24" )
   END_RUNG wire#w2
   // the same network as SCL:
   "DB_GENERAL".Concatenadoras[12] := "DB_GENERAL".Estados[11] AND (#DoneYN OR "Band_E24") AND "DB_GENERAL".Cuenta_3 AND NOT "DB_INC_GENERAL".Alarma_On;
END_REGION

REGION Network 23: Concatenadora 13
   RUNG wire#powerrail
      Contact( "DB_GENERAL".Estados[12] )
      Contact( #DoneXN )
      Contact( #DoneY )
      wire#w1
      I_Contact( "DB_INC_GENERAL".Alarma_On )
      Coil( "DB_GENERAL".Concatenadoras[13] )
   END_RUNG
   RUNG wire#powerrail
      Contact( "DB_GENERAL".Estados[23] )
      I_Contact( "01_LINEA_Entradas-DB".Canal3_Full )
      Contact( "01_LINEA_Entradas-DB".Canal1_Full )
   END_RUNG wire#w1
   // the same network as SCL:
   "DB_GENERAL".Concatenadoras[13] := (("DB_GENERAL".Estados[12] AND #DoneXN AND #DoneY) OR ("DB_GENERAL".Estados[23] AND NOT "01_LINEA_Entradas-DB".Canal3_Full AND "01_LINEA_Entradas-DB".Canal1_Full)) AND NOT "DB_INC_GENERAL".Alarma_On;
END_REGION

REGION Network 24: Concatenadora 14
   RUNG wire#powerrail
      Contact( "DB_GENERAL".Estados[13] )
      wire#w1
      Contact( #DoneYN )
      wire#w2
      Contact( "DB_GENERAL".Cuenta_1 )
      I_Contact( "DB_INC_GENERAL".Alarma_On )
      Coil( "DB_GENERAL".Concatenadoras[10] )
   END_RUNG
   RUNG wire#w1
      Contact( "Band_E23" )
   END_RUNG wire#w2
   // the same network as SCL:
   "DB_GENERAL".Concatenadoras[10] := "DB_GENERAL".Estados[13] AND (#DoneYN OR "Band_E23") AND "DB_GENERAL".Cuenta_1 AND NOT "DB_INC_GENERAL".Alarma_On;
END_REGION

REGION Network 25: Concatenadora 15
   RUNG wire#powerrail
      Contact( "DB_GENERAL".Estados[14] )
      wire#w1
      Contact( #Done2X )
      wire#w2
      Contact( #DoneY )
      wire#w3
      I_Contact( "DB_INC_GENERAL".Alarma_On )
      Coil( "DB_GENERAL".Concatenadoras[15] )
   END_RUNG
   RUNG wire#w1
      Contact( #DoneX )
   END_RUNG wire#w2
   RUNG wire#powerrail
      Contact( "DB_GENERAL".Estados[24] )
      I_Contact( "01_LINEA_Entradas-DB".Canal1_Full )
      Contact( "01_LINEA_Entradas-DB".Canal2_Full )
   END_RUNG wire#w3
   // the same network as SCL:
   "DB_GENERAL".Concatenadoras[15] := (("DB_GENERAL".Estados[14] AND (#Done2X OR #DoneX) AND #DoneY) OR ("DB_GENERAL".Estados[24] AND NOT "01_LINEA_Entradas-DB".Canal1_Full AND "01_LINEA_Entradas-DB".Canal2_Full)) AND NOT "DB_INC_GENERAL".Alarma_On;
END_REGION

REGION Network 26: Concatenadora 16
   RUNG wire#powerrail
      Contact( "DB_GENERAL".Estados[15] )
      wire#w1
      Contact( #DoneYN )
      wire#w2
      Contact( "DB_GENERAL".Cuenta_3 )
      I_Contact( "DB_INC_GENERAL".Alarma_On )
      Coil( "DB_GENERAL".Concatenadoras[16] )
   END_RUNG
   RUNG wire#w1
      Contact( "Band_E24" )
   END_RUNG wire#w2
   // the same network as SCL:
   "DB_GENERAL".Concatenadoras[16] := "DB_GENERAL".Estados[15] AND (#DoneYN OR "Band_E24") AND "DB_GENERAL".Cuenta_3 AND NOT "DB_INC_GENERAL".Alarma_On;
END_REGION

REGION Network 27: Concatenadora 17
   RUNG wire#powerrail
      Contact( "DB_GENERAL".Estados[16] )
      Contact( #Done2XN )
      Contact( #DoneY )
      wire#w1
      I_Contact( "DB_INC_GENERAL".Alarma_On )
      Coil( "DB_GENERAL".Concatenadoras[17] )
   END_RUNG
   RUNG wire#powerrail
      Contact( "DB_GENERAL".Estados[22] )
      I_Contact( "01_LINEA_Entradas-DB".Canal3_Full )
      Contact( "01_LINEA_Entradas-DB".Canal2_Full )
   END_RUNG wire#w1
   // the same network as SCL:
   "DB_GENERAL".Concatenadoras[17] := (("DB_GENERAL".Estados[16] AND #Done2XN AND #DoneY) OR ("DB_GENERAL".Estados[22] AND NOT "01_LINEA_Entradas-DB".Canal3_Full AND "01_LINEA_Entradas-DB".Canal2_Full)) AND NOT "DB_INC_GENERAL".Alarma_On;
END_REGION

REGION Network 28: Concatenadora 18
   RUNG wire#powerrail
      Contact( "DB_GENERAL".Estados[17] )
      wire#w1
      Contact( #DoneYN )
      wire#w2
      Contact( "DB_GENERAL".Cuenta_1 )
      I_Contact( "DB_INC_GENERAL".Alarma_On )
      Coil( "DB_GENERAL".Concatenadoras[14] )
   END_RUNG
   RUNG wire#w1
      Contact( "Band_E22" )
   END_RUNG wire#w2
   // the same network as SCL:
   "DB_GENERAL".Concatenadoras[14] := "DB_GENERAL".Estados[17] AND (#DoneYN OR "Band_E22") AND "DB_GENERAL".Cuenta_1 AND NOT "DB_INC_GENERAL".Alarma_On;
END_REGION

REGION Network 29: Concatenadora 19